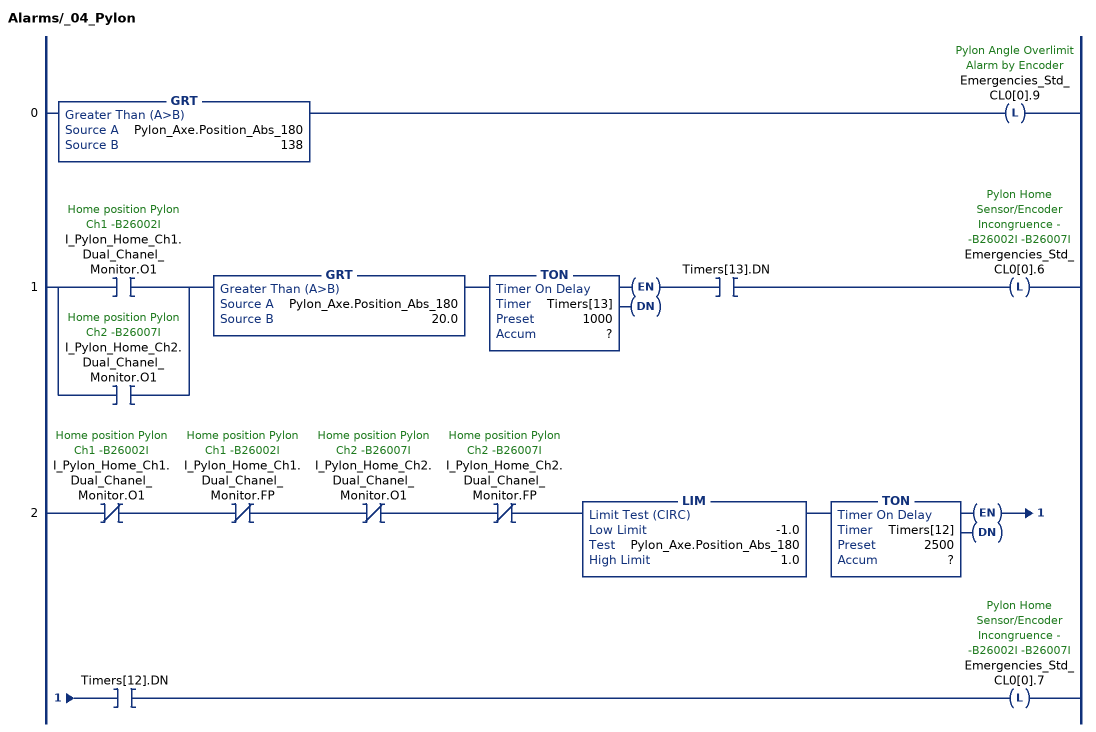
   0: GRT(Pylon_Axe.Position_Abs_180,138)OTL(Emergencies_Std_CL0[0].9);
   1: [XIC(I_Pylon_Home_Ch1.Dual_Chanel_Monitor.O1) ,XIC(I_Pylon_Home_Ch2.Dual_Chanel_Monitor.O1) ]GRT(Pylon_Axe.Position_Abs_180,20.0)TON(Timers[13],?,?)XIC(Timers[13].DN)OTL(Emergencies_Std_CL0[0].6);
   2: XIO(I_Pylon_Home_Ch1.Dual_Chanel_Monitor.O1)XIO(I_Pylon_Home_Ch1.Dual_Chanel_Monitor.FP)XIO(I_Pylon_Home_Ch2.Dual_Chanel_Monitor.O1)XIO(I_Pylon_Home_Ch2.Dual_Chanel_Monitor.FP)LIM(-1.0,Pylon_Axe.Position_Abs_180,1.0)TON(Timers[12],?,?)XIC(Timers[12].DN)OTL(Emergencies_Std_CL0[0].7);
END_ROUTINE

ROUTINE Main   (* ladder *)
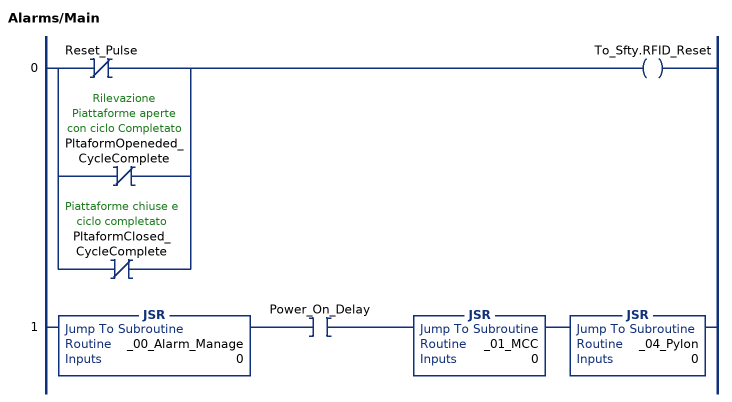
   0: [XIO(Reset_Pulse) ,XIO(PltaformOpeneded_CycleComplete) ,XIO(PltaformClosed_CycleComplete) ]OTE(To_Sfty.RFID_Reset);
   1: JSR(_00_Alarm_Manage,0)XIC(Power_On_Delay)JSR(_01_MCC,0)JSR(_04_Pylon,0);
END_ROUTINE
END_PROGRAM

PROGRAM General   (* main routine Main *)
VAR
   Avg_TimeInStation_CurrentHour : DINT := 303;
   Avg_TimeInStation_Daily : DINT := 207;
   Closing_CyclePlatTimes : DINT[20] := ([1] := 60000, [2] := 679, [3] := 679, [4] := 17399, [5] := 19639, [6] := 19639, [9] := 16239, [10] := 3400);
        [14]   // daily avg overall
        [13]   // daily total overall
        [11]   // daily total time waiting
        [10]   // Time Waiting on Lever,etc
        [9]   // Time Platform Move In Close
        [12]   // daily avg time waiting
   Cycle_Before_Timer : TIMER := (PRE := 60000);
   CyclePlatClose_Count_Daily : COUNTER := (PRE := 500);
   CyclePlatOpen_Count_Daily : COUNTER := (PRE := 500);
   DAY : DINT := 1;   // Day
   HMI_LapBars_Status : DINT := 1;   // 0 = Closed 1 = Opened 2 = Closing 3 = Opening
   HMI_Platform_Status : DINT := 1;   // 0 = Stopped 1 = Closing 2 = Closed 3 = Opening 4 = Opened
   HMI_reset_Partial_Life_Cycle : BOOL;
   HMI_reset_Partial_Life_RunHH : BOOL;
   HOUR : DINT := 19;   // Hour
   JM_Statistics_Hist : Run_Count_Hist_JM[100] := ([0].date[0] := 25, [0].date[1] := 11, [0].date[2] := 29, [0].runs[0] := 11, [0].runs[7] := 1, [0].runs[8] := 2, [0].runs[9] := 2, [0].runs[13] := 4, [0].runs[15] := 1, [0].runs[19] := 3, [0].time_avg[0] := 207, [0].time_avg[4] := 19639, [0].time_avg[5] := 22361, [0].time_avg[8] := 48, [0].time_avg[9] := 48, [0].time_avg[13] := 196, [0].time_avg[19] := 303, [1].date[0] := 25, [1].date[1] := 11, [1].date[2] := 28, [1].runs[0] := 65, [1].runs[8] := 2, [1].runs[9] := 1, [1].runs[15] := 3, [1].runs[16] := 7, [1].runs[17] := 8, [1].runs[18] := 8, [1].runs[19] := 8, [1].runs[20] := 8, [1].runs[21] := 7, [1].runs[22] := 8, [1].runs[23] := 5, [1].time_avg[0] := 204, [1].time_avg[2] := 3400, [1].time_avg[4] := 19639, [1].time_avg[5] := 22361, [1].time_avg[8] := 50, [1].time_avg[15] := 203, [1].time_avg[16] := 254, [1].time_avg[17] := 210, [1].time_avg[18] := 202, [1].time_avg[19] := 195, [1].time_avg[20] := 206, [1].time_avg[21] := 190, [1].time_avg[22] := 211, [1].time_avg[23] := 177, [2].date[0] := 25, [2].date[1] := 11, [2].date[2] := 27, [2].runs[0] := 63, [2].runs[14] := 6, [2].runs[15] := 4, [2].runs[16] := 7, [2].runs[17] := 7, [2].runs[18] := 8, [2].runs[19] := 8, [2].runs[20] := 7, [2].runs[21] := 5, [2].runs[22] := 8, [2].runs[23] := 3,
        [2].time_avg[0] := 234, [2].time_avg[4] := 21760, [2].time_avg[5] := 22361, [2].time_avg[14] := 167, [2].time_avg[15] := 316, [2].time_avg[16] := 272, [2].time_avg[17] := 206, [2].time_avg[18] := 208, [2].time_avg[19] := 242, [2].time_avg[20] := 266, [2].time_avg[21] := 233, [2].time_avg[22] := 223, [2].time_avg[23] := 245, [3].date[0] := 25, [3].date[1] := 11, [3].date[2] := 26, [3].runs[0] := 57, [3].runs[12] := 4, [3].runs[13] := 1, [3].runs[15] := 2, [3].runs[16] := 6, [3].runs[17] := 7, [3].runs[18] := 7, [3].runs[19] := 7, [3].runs[20] := 7, [3].runs[21] := 7, [3].runs[22] := 6, [3].runs[23] := 3, [3].time_avg[0] := 274, [3].time_avg[2] := 6041, [3].time_avg[4] := 21760, [3].time_avg[5] := 22361, [3].time_avg[12] := 396, [3].time_avg[13] := 320, [3].time_avg[15] := 271, [3].time_avg[16] := 271, [3].time_avg[17] := 292, [3].time_avg[18] := 243, [3].time_avg[19] := 255, [3].time_avg[20] := 243, [3].time_avg[21] := 289, [3].time_avg[22] := 278, [3].time_avg[23] := 283, [4].date[0] := 25, [4].date[1] := 11, [4].date[2] := 25, [4].runs[0] := 53, [4].runs[7] := 1, [4].runs[15] := 1, [4].runs[16] := 5, [4].runs[17] := 8, [4].runs[18] := 6, [4].runs[19] := 8, [4].runs[20] := 7, [4].runs[21] := 7, [4].runs[22] := 7, [4].runs[23] := 3, [4].time_avg[0] := 260, [4].time_avg[4] := 53080, [4].time_avg[5] := 22361,
        [4].time_avg[16] := 223, [4].time_avg[17] := 286, [4].time_avg[18] := 280, [4].time_avg[19] := 258, [4].time_avg[20] := 261, [4].time_avg[21] := 234, [4].time_avg[22] := 267, [4].time_avg[23] := 254, [5].date[0] := 25, [5].date[1] := 11, [5].date[2] := 24, [5].runs[0] := 67, [5].runs[7] := 4, [5].runs[8] := 3, [5].runs[10] := 2, [5].runs[11] := 4, [5].runs[13] := 1, [5].runs[14] := 1, [5].runs[15] := 4, [5].runs[16] := 7, [5].runs[17] := 7, [5].runs[18] := 7, [5].runs[19] := 7, [5].runs[20] := 4, [5].runs[21] := 7, [5].runs[22] := 6, [5].runs[23] := 3, [5].time_avg[0] := 254, [5].time_avg[2] := 76642, [5].time_avg[4] := 53080, [5].time_avg[5] := 22361, [5].time_avg[7] := 75, [5].time_avg[8] := 246, [5].time_avg[11] := 171, [5].time_avg[14] := 83, [5].time_avg[15] := 147, [5].time_avg[16] := 272, [5].time_avg[17] := 276, [5].time_avg[18] := 244, [5].time_avg[19] := 256, [5].time_avg[20] := 266, [5].time_avg[21] := 291, [5].time_avg[22] := 291, [5].time_avg[23] := 290, [6].date[0] := 25, [6].date[1] := 11, [6].date[2] := 23, [6].runs[0] := 54, [6].runs[10] := 2, [6].runs[11] := 4, [6].runs[15] := 1, [6].runs[16] := 8, [6].runs[17] := 7, [6].runs[18] := 6, [6].runs[19] := 5, [6].runs[20] := 8, [6].runs[21] := 6, [6].runs[22] := 5, [6].runs[23] := 2, [6].time_avg[0] := 268,
        [6].time_avg[4] := 23760, [6].time_avg[5] := 22361, [6].time_avg[11] := 332, [6].time_avg[16] := 211, [6].time_avg[17] := 253, [6].time_avg[18] := 262, [6].time_avg[19] := 274, [6].time_avg[20] := 241, [6].time_avg[21] := 295, [6].time_avg[22] := 310, [6].time_avg[23] := 371, [7].date[0] := 25, [7].date[1] := 11, [7].date[2] := 22, [7].runs[0] := 49, [7].runs[12] := 7, [7].runs[14] := 1, [7].runs[15] := 4, [7].runs[16] := 7, [7].runs[17] := 7, [7].runs[18] := 7, [7].runs[19] := 1, [7].runs[20] := 6, [7].runs[21] := 2, [7].runs[22] := 6, [7].runs[23] := 1, [7].time_avg[0] := 278, [7].time_avg[4] := 23760, [7].time_avg[5] := 22361, [7].time_avg[12] := 180, [7].time_avg[15] := 308, [7].time_avg[16] := 282, [7].time_avg[17] := 261, [7].time_avg[18] := 280, [7].time_avg[19] := 295, [7].time_avg[20] := 361, [7].time_avg[22] := 287, [8].date[0] := 25, [8].date[1] := 11, [8].date[2] := 20, [8].runs[0] := 58, [8].runs[10] := 2, [8].runs[11] := 3, [8].runs[13] := 5, [8].runs[14] := 4, [8].runs[15] := 3, [8].runs[16] := 5, [8].runs[17] := 4, [8].runs[18] := 3, [8].runs[19] := 6, [8].runs[20] := 5, [8].runs[21] := 7, [8].runs[22] := 7, [8].runs[23] := 4, [8].time_avg[0] := 205, [8].time_avg[2] := 15381, [8].time_avg[4] := 23760, [8].time_avg[5] := 22361, [8].time_avg[10] := 76, [8].time_avg[11] := 152,
        [8].time_avg[13] := 198, [8].time_avg[14] := 60, [8].time_avg[15] := 73, [8].time_avg[16] := 76, [8].time_avg[17] := 183, [8].time_avg[18] := 376, [8].time_avg[19] := 286, [8].time_avg[20] := 250, [8].time_avg[21] := 218, [8].time_avg[22] := 239, [8].time_avg[23] := 211, [9].date[0] := 25, [9].date[1] := 11, [9].date[2] := 19, [9].runs[0] := 7, [9].runs[12] := 2, [9].runs[13] := 4, [9].runs[17] := 1, [9].runs[18] := 1, [9].time_avg[0] := 217, [9].time_avg[2] := 78801, [9].time_avg[4] := 48480, [9].time_avg[5] := 22361, [9].time_avg[13] := 217, [10].date[0] := 25, [10].date[1] := 11, [10].date[2] := 16, [10].runs[0] := 7, [10].runs[10] := 2, [10].runs[13] := 7, [10].time_avg[0] := 93, [10].time_avg[4] := 27759, [10].time_avg[5] := 22361, [10].time_avg[13] := 93, [11].date[0] := 25, [11].date[1] := 11, [11].date[2] := 14, [11].runs[0] := 2, [11].runs[15] := 1, [11].runs[16] := 1, [11].time_avg[2] := 32760, [11].time_avg[4] := 27759, [11].time_avg[5] := 22361, [12].date[0] := 25, [12].date[1] := 11, [12].date[2] := 13, [12].runs[0] := 14, [12].runs[10] := 2, [12].runs[11] := 1, [12].runs[12] := 1, [12].runs[14] := 2, [12].runs[15] := 5, [12].runs[16] := 4, [12].runs[17] := 5, [12].time_avg[0] := 141, [12].time_avg[4] := 36240, [12].time_avg[5] := 22361, [12].time_avg[10] := 210, [12].time_avg[14] := 205, [12].time_avg[15] := 160,
        [12].time_avg[16] := 100, [12].time_avg[17] := 100, [13].date[0] := 25, [13].date[1] := 11, [13].date[2] := 11, [13].runs[0] := 2, [13].runs[18] := 2, [13].time_avg[0] := 88, [13].time_avg[4] := 36240, [13].time_avg[5] := 22361, [13].time_avg[18] := 88, [14].date[0] := 25, [14].date[1] := 11, [14].date[2] := 7, [14].runs[0] := 5, [14].runs[15] := 3, [14].runs[16] := 2, [14].time_avg[0] := 229, [14].time_avg[4] := 36240, [14].time_avg[5] := 22361, [14].time_avg[15] := 300, [14].time_avg[16] := 87, [15].date[0] := 25, [15].date[1] := 11, [15].date[2] := 6, [15].runs[0] := 13, [15].runs[15] := 1, [15].runs[16] := 3, [15].runs[17] := 8, [15].runs[18] := 1, [15].runs[19] := 4, [15].time_avg[0] := 54, [15].time_avg[4] := 36240, [15].time_avg[5] := 22361, [15].time_avg[17] := 46, [15].time_avg[19] := 66, [16].date[0] := 25, [16].date[1] := 10, [16].date[2] := 27, [16].runs[0] := 13, [16].runs[12] := 1, [16].runs[13] := 4, [16].runs[14] := 1, [16].time_avg[0] := 126, [16].time_avg[4] := 36240, [16].time_avg[5] := 22361, [16].time_avg[13] := 65, [17].date[0] := 25, [17].date[1] := 10, [17].date[2] := 26, [17].runs[0] := 58, [17].runs[10] := 1, [17].runs[11] := 2, [17].runs[12] := 3, [17].runs[13] := 8, [17].runs[14] := 8, [17].runs[15] := 6, [17].runs[16] := 7, [17].runs[17] := 7, [17].runs[18] := 6,
        [17].runs[19] := 7, [17].runs[20] := 3, [17].time_avg[0] := 252, [17].time_avg[2] := 40720, [17].time_avg[4] := 36240, [17].time_avg[5] := 22361, [17].time_avg[11] := 476, [17].time_avg[12] := 190, [17].time_avg[13] := 206, [17].time_avg[14] := 216, [17].time_avg[15] := 310, [17].time_avg[16] := 261, [17].time_avg[17] := 248, [17].time_avg[18] := 232, [17].time_avg[19] := 304, [17].time_avg[20] := 214, [18].date[0] := 25, [18].date[1] := 10, [18].date[2] := 25, [18].runs[0] := 47, [18].runs[12] := 5, [18].runs[13] := 9, [18].runs[14] := 5, [18].runs[16] := 2, [18].runs[17] := 8, [18].runs[18] := 7, [18].runs[19] := 7, [18].runs[20] := 4, [18].time_avg[0] := 227, [18].time_avg[4] := 26040, [18].time_avg[5] := 22361, [18].time_avg[12] := 203, [18].time_avg[13] := 166, [18].time_avg[14] := 231, [18].time_avg[16] := 370, [18].time_avg[17] := 239, [18].time_avg[18] := 252, [18].time_avg[19] := 244, [18].time_avg[20] := 235, [19].date[0] := 25, [19].date[1] := 10, [19].date[2] := 23, [19].runs[0] := 48, [19].runs[9] := 2, [19].runs[10] := 3, [19].runs[12] := 3, [19].runs[13] := 7, [19].runs[14] := 7, [19].runs[15] := 5, [19].runs[16] := 8, [19].runs[17] := 5, [19].runs[19] := 5, [19].runs[20] := 3, [19].time_avg[0] := 257, [19].time_avg[2] := 18201, [19].time_avg[4] := 26040, [19].time_avg[5] := 22361, [19].time_avg[9] := 102, [19].time_avg[10] := 259, [19].time_avg[12] := 493,
        [19].time_avg[13] := 241, [19].time_avg[14] := 231, [19].time_avg[15] := 264, [19].time_avg[16] := 252, [19].time_avg[17] := 280, [19].time_avg[19] := 300, [19].time_avg[20] := 235, [20].date[0] := 25, [20].date[1] := 10, [20].date[2] := 22, [20].runs[0] := 62, [20].runs[10] := 4, [20].runs[12] := 2, [20].runs[13] := 9, [20].runs[14] := 7, [20].runs[15] := 7, [20].runs[16] := 7, [20].runs[17] := 7, [20].runs[18] := 8, [20].runs[19] := 8, [20].runs[20] := 3, [20].time_avg[0] := 226, [20].time_avg[4] := 26079, [20].time_avg[5] := 22361, [20].time_avg[10] := 123, [20].time_avg[13] := 199, [20].time_avg[14] := 230, [20].time_avg[15] := 230, [20].time_avg[16] := 312, [20].time_avg[17] := 253, [20].time_avg[18] := 219, [20].time_avg[19] := 200, [20].time_avg[20] := 206, [21].date[0] := 25, [21].date[1] := 10, [21].date[2] := 21, [21].runs[0] := 58, [21].runs[11] := 3, [21].runs[12] := 1, [21].runs[13] := 8, [21].runs[14] := 7, [21].runs[15] := 4, [21].runs[16] := 8, [21].runs[17] := 8, [21].runs[18] := 7, [21].runs[19] := 8, [21].runs[20] := 4, [21].time_avg[0] := 233, [21].time_avg[2] := 42160, [21].time_avg[4] := 26079, [21].time_avg[5] := 22361, [21].time_avg[11] := 186, [21].time_avg[13] := 222, [21].time_avg[14] := 240, [21].time_avg[15] := 294, [21].time_avg[16] := 256, [21].time_avg[17] := 202, [21].time_avg[18] := 246, [21].time_avg[19] := 216, [21].time_avg[20] := 208,
        [22].date[0] := 25, [22].date[1] := 10, [22].date[2] := 20, [22].runs[0] := 47, [22].runs[10] := 2, [22].runs[11] := 6, [22].runs[12] := 1, [22].runs[13] := 7, [22].runs[14] := 7, [22].runs[15] := 7, [22].runs[16] := 4, [22].runs[17] := 1, [22].runs[18] := 2, [22].runs[19] := 7, [22].runs[20] := 3, [22].time_avg[0] := 249, [22].time_avg[2] := 52640, [22].time_avg[4] := 40960, [22].time_avg[5] := 22361, [22].time_avg[11] := 232, [22].time_avg[13] := 215, [22].time_avg[14] := 258, [22].time_avg[15] := 237, [22].time_avg[16] := 210, [22].time_avg[18] := 331, [22].time_avg[19] := 294, [22].time_avg[20] := 241, [23].date[0] := 25, [23].date[1] := 10, [23].date[2] := 19, [23].runs[0] := 61, [23].runs[9] := 2, [23].runs[10] := 2, [23].runs[11] := 8, [23].runs[12] := 4, [23].runs[13] := 6, [23].runs[14] := 1, [23].runs[15] := 8, [23].runs[16] := 7, [23].runs[17] := 7, [23].runs[18] := 7, [23].runs[19] := 7, [23].runs[20] := 2, [23].time_avg[0] := 237, [23].time_avg[2] := 59762, [23].time_avg[4] := 52320, [23].time_avg[5] := 22361, [23].time_avg[9] := 89, [23].time_avg[11] := 203, [23].time_avg[12] := 193, [23].time_avg[13] := 194, [23].time_avg[15] := 243, [23].time_avg[16] := 238, [23].time_avg[17] := 251, [23].time_avg[18] := 268, [23].time_avg[19] := 280, [23].time_avg[20] := 287, [24].date[0] := 25, [24].date[1] := 10, [24].date[2] := 18,
        [24].runs[0] := 51, [24].runs[9] := 2, [24].runs[10] := 5, [24].runs[11] := 8, [24].runs[12] := 2, [24].runs[13] := 5, [24].runs[14] := 6, [24].runs[15] := 7, [24].runs[16] := 5, [24].runs[17] := 7, [24].runs[18] := 4, [24].time_avg[0] := 246, [24].time_avg[4] := 52360, [24].time_avg[5] := 22361, [24].time_avg[10] := 182, [24].time_avg[11] := 228, [24].time_avg[12] := 212, [24].time_avg[13] := 231, [24].time_avg[14] := 324, [24].time_avg[15] := 255, [24].time_avg[16] := 238, [24].time_avg[17] := 263, [24].time_avg[18] := 255, [25].date[0] := 25, [25].date[1] := 10, [25].date[2] := 15, [25].runs[0] := 89, [25].runs[10] := 4, [25].runs[11] := 4, [25].runs[12] := 7, [25].runs[13] := 6, [25].runs[14] := 8, [25].runs[15] := 6, [25].runs[16] := 7, [25].runs[17] := 6, [25].time_avg[0] := 251, [25].time_avg[2] := 50482, [25].time_avg[4] := 52360, [25].time_avg[5] := 22361, [25].time_avg[10] := 61, [25].time_avg[11] := 214, [25].time_avg[12] := 261, [25].time_avg[13] := 348, [25].time_avg[14] := 197, [25].time_avg[15] := 264, [25].time_avg[16] := 241, [25].time_avg[17] := 309, [26].date[0] := 25, [26].date[1] := 10, [26].date[2] := 14, [26].runs[0] := 14, [26].runs[10] := 5, [26].runs[11] := 1, [26].runs[12] := 8, [26].time_avg[0] := 175, [26].time_avg[4] := 34119, [26].time_avg[5] := 22361, [26].time_avg[10] := 270, [26].time_avg[12] := 121, [27].date[0] := 25,
        [27].date[1] := 10, [27].date[2] := 13, [27].runs[0] := 29, [27].runs[12] := 3, [27].runs[13] := 5, [27].runs[14] := 6, [27].runs[15] := 4, [27].runs[16] := 7, [27].runs[17] := 4, [27].time_avg[0] := 256, [27].time_avg[2] := 63880, [27].time_avg[4] := 34119, [27].time_avg[5] := 22361, [27].time_avg[12] := 68, [27].time_avg[13] := 218, [27].time_avg[14] := 246, [27].time_avg[15] := 367, [27].time_avg[16] := 315, [27].time_avg[17] := 255, [28].date[0] := 25, [28].date[1] := 10, [28].date[2] := 10, [28].runs[0] := 27, [28].runs[9] := 9, [28].runs[10] := 11, [28].runs[11] := 7, [28].time_avg[0] := 89, [28].time_avg[4] := 33481, [28].time_avg[5] := 22361, [28].time_avg[9] := 82, [28].time_avg[10] := 83, [28].time_avg[11] := 123, [29].date[0] := 25, [29].date[1] := 10, [29].date[2] := 8, [29].runs[0] := 76, [29].runs[9] := 9, [29].runs[10] := 11, [29].runs[11] := 8, [29].runs[12] := 10, [29].runs[13] := 11, [29].runs[14] := 7, [29].runs[15] := 7, [29].runs[16] := 3, [29].time_avg[0] := 100, [29].time_avg[4] := 33481, [29].time_avg[5] := 22361, [29].time_avg[9] := 47, [29].time_avg[10] := 77, [29].time_avg[11] := 96, [29].time_avg[12] := 96, [29].time_avg[13] := 82, [29].time_avg[14] := 70, [29].time_avg[15] := 221, [29].time_avg[16] := 56, [30].date[0] := 25, [30].date[1] := 10, [30].date[2] := 7, [30].runs[0] := 1, [30].runs[8] := 1,
        [30].time_avg[4] := 33481, [30].time_avg[5] := 22361, [31].date[0] := 25, [31].date[1] := 10, [31].date[2] := 6, [31].runs[0] := 3, [31].runs[12] := 3, [31].time_avg[0] := 51, [31].time_avg[4] := 33481, [31].time_avg[5] := 22361, [31].time_avg[12] := 51, [32].date[0] := 25, [32].date[1] := 10, [32].date[2] := 5, [32].runs[0] := 3, [32].runs[12] := 1, [32].runs[15] := 2, [32].time_avg[0] := 43, [32].time_avg[4] := 33481, [32].time_avg[5] := 22361, [32].time_avg[15] := 43, [33].date[0] := 25, [33].date[1] := 10, [33].date[2] := 4, [33].runs[0] := 15, [33].runs[10] := 4, [33].runs[11] := 3, [33].runs[12] := 3, [33].runs[15] := 4, [33].runs[16] := 1, [33].time_avg[0] := 228, [33].time_avg[2] := 47342, [33].time_avg[4] := 33481, [33].time_avg[5] := 22361, [33].time_avg[10] := 258, [33].time_avg[11] := 342, [33].time_avg[12] := 69, [33].time_avg[15] := 112, [34].date[0] := 25, [34].date[1] := 10, [34].date[2] := 1, [34].runs[0] := 64, [34].runs[9] := 1, [34].runs[10] := 7, [34].runs[11] := 8, [34].runs[12] := 9, [34].runs[13] := 6, [34].runs[14] := 8, [34].runs[15] := 9, [34].runs[16] := 8, [34].runs[17] := 8, [34].time_avg[0] := 168, [34].time_avg[4] := 53200, [34].time_avg[5] := 22361, [34].time_avg[10] := 151, [34].time_avg[11] := 172, [34].time_avg[12] := 168, [34].time_avg[13] := 171, [34].time_avg[14] := 150, [34].time_avg[15] := 177,
        [34].time_avg[16] := 175, [34].time_avg[17] := 175, [35].date[0] := 25, [35].date[1] := 9, [35].date[2] := 30, [35].runs[0] := 60, [35].runs[9] := 5, [35].runs[10] := 5, [35].runs[11] := 9, [35].runs[12] := 7, [35].runs[13] := 8, [35].runs[14] := 9, [35].runs[15] := 9, [35].runs[16] := 8, [35].time_avg[0] := 176, [35].time_avg[2] := 40561, [35].time_avg[4] := 53200, [35].time_avg[5] := 22361, [35].time_avg[9] := 120, [35].time_avg[10] := 150, [35].time_avg[11] := 176, [35].time_avg[12] := 186, [35].time_avg[13] := 219, [35].time_avg[14] := 153, [35].time_avg[15] := 180, [35].time_avg[16] := 165, [36].date[0] := 25, [36].date[1] := 9, [36].date[2] := 29, [36].runs[0] := 57, [36].runs[8] := 2, [36].runs[9] := 7, [36].runs[10] := 7, [36].runs[11] := 8, [36].runs[12] := 5, [36].runs[13] := 7, [36].runs[14] := 7, [36].runs[15] := 7, [36].runs[16] := 7, [36].time_avg[0] := 211, [36].time_avg[4] := 56839, [36].time_avg[5] := 22361, [36].time_avg[9] := 166, [36].time_avg[10] := 267, [36].time_avg[11] := 147, [36].time_avg[12] := 241, [36].time_avg[13] := 205, [36].time_avg[14] := 168, [36].time_avg[15] := 266, [36].time_avg[16] := 222, [37].date[0] := 25, [37].date[1] := 9, [37].date[2] := 28, [37].runs[0] := 58, [37].runs[9] := 3, [37].runs[10] := 9, [37].runs[11] := 7, [37].runs[12] := 8, [37].runs[13] := 8, [37].runs[14] := 8,
        [37].runs[15] := 7, [37].runs[16] := 8, [37].time_avg[0] := 184, [37].time_avg[4] := 56839, [37].time_avg[5] := 22361, [37].time_avg[9] := 167, [37].time_avg[10] := 193, [37].time_avg[11] := 208, [37].time_avg[12] := 169, [37].time_avg[13] := 199, [37].time_avg[14] := 199, [37].time_avg[15] := 173, [37].time_avg[16] := 151, [38].date[0] := 25, [38].date[1] := 9, [38].date[2] := 25, [38].runs[0] := 64, [38].runs[8] := 4, [38].runs[9] := 6, [38].runs[10] := 7, [38].runs[11] := 7, [38].runs[12] := 8, [38].runs[13] := 8, [38].runs[14] := 8, [38].runs[15] := 9, [38].runs[16] := 7, [38].time_avg[0] := 201, [38].time_avg[4] := 56839, [38].time_avg[5] := 22361, [38].time_avg[8] := 455, [38].time_avg[9] := 193, [38].time_avg[10] := 212, [38].time_avg[11] := 189, [38].time_avg[12] := 207, [38].time_avg[13] := 224, [38].time_avg[14] := 191, [38].time_avg[15] := 166, [38].time_avg[16] := 193, [39].date[0] := 25, [39].date[1] := 9, [39].date[2] := 24, [39].runs[0] := 50, [39].runs[9] := 4, [39].runs[10] := 6, [39].runs[11] := 5, [39].runs[12] := 6, [39].runs[13] := 5, [39].runs[14] := 8, [39].runs[15] := 8, [39].runs[16] := 8, [39].time_avg[0] := 195, [39].time_avg[4] := 56839, [39].time_avg[5] := 22361, [39].time_avg[9] := 83, [39].time_avg[10] := 198, [39].time_avg[11] := 260, [39].time_avg[12] := 133, [39].time_avg[13] := 207, [39].time_avg[14] := 244, [39].time_avg[15] := 215,
        [39].time_avg[16] := 169, [40].date[0] := 25, [40].date[1] := 9, [40].date[2] := 22, [40].runs[0] := 46, [40].runs[8] := 4, [40].runs[9] := 3, [40].runs[10] := 7, [40].runs[11] := 5, [40].runs[12] := 7, [40].runs[13] := 5, [40].runs[14] := 2, [40].runs[15] := 6, [40].runs[16] := 7, [40].time_avg[0] := 229, [40].time_avg[4] := 56839, [40].time_avg[5] := 22361, [40].time_avg[8] := 208, [40].time_avg[10] := 179, [40].time_avg[11] := 196, [40].time_avg[12] := 160, [40].time_avg[13] := 227, [40].time_avg[15] := 325, [40].time_avg[16] := 281, [41].date[0] := 25, [41].date[1] := 9, [41].date[2] := 21, [41].runs[0] := 9, [41].runs[8] := 1, [41].runs[9] := 6, [41].runs[14] := 2, [41].time_avg[0] := 233, [41].time_avg[2] := 43360, [41].time_avg[4] := 56839, [41].time_avg[5] := 22361, [41].time_avg[9] := 244, [41].time_avg[14] := 175, [42].date[0] := 25, [42].date[1] := 9, [42].date[2] := 18, [42].runs[0] := 6, [42].runs[11] := 5, [42].runs[12] := 1, [42].time_avg[0] := 226, [42].time_avg[4] := 37320, [42].time_avg[5] := 22361, [42].time_avg[11] := 226, [43].date[0] := 25, [43].date[1] := 9, [43].date[2] := 16, [43].runs[0] := 2, [43].runs[15] := 1, [43].runs[16] := 1, [43].time_avg[2] := 46801, [43].time_avg[4] := 37320, [43].time_avg[5] := 22361, [44].date[0] := 25, [44].date[1] := 8, [44].date[2] := 15, [44].runs[0] := 3,
        [44].runs[12] := 1, [44].runs[15] := 2, [44].time_avg[4] := 37641, [44].time_avg[5] := 22361, [45].date[0] := 25, [45].date[1] := 7, [45].date[2] := 13, [45].runs[0] := 107, [45].runs[9] := 2, [45].runs[14] := 2, [45].runs[16] := 8, [45].time_avg[0] := 162, [45].time_avg[2] := 22208, [45].time_avg[4] := 37641, [45].time_avg[5] := 22361, [45].time_avg[9] := 55, [45].time_avg[14] := 220, [45].time_avg[16] := 142, [46].date[0] := -2, [46].date[1] := 1, [46].date[2] := 15, [46].runs[0] := 1, [46].time_avg[4] := 45599, [46].time_avg[5] := 22361, [47].date[0] := -2, [47].date[1] := 1, [47].date[2] := 12, [47].runs[0] := 14, [47].runs[23] := 3, [47].time_avg[0] := 172, [47].time_avg[4] := 45599, [47].time_avg[5] := 22361, [47].time_avg[23] := 108, [48].date[0] := -2, [48].date[1] := 1, [48].date[2] := 11, [48].runs[0] := 14, [48].runs[21] := 1, [48].time_avg[0] := 145, [48].time_avg[4] := 45599, [48].time_avg[5] := 22361, [49].date[0] := -2, [49].date[1] := 1, [49].date[2] := 10, [49].runs[0] := 2, [49].runs[20] := 1, [49].runs[23] := 1, [49].time_avg[4] := 45599, [49].time_avg[5] := 22361, [50].date[0] := -2, [50].date[1] := 1, [50].date[2] := 8, [50].runs[0] := 1, [50].time_avg[4] := 45599, [50].time_avg[5] := 22361, [51].date[0] := -2, [51].date[1] := 1, [51].date[2] := 6, [51].runs[0] := 2, [51].runs[20] := 1,
        [51].time_avg[4] := 45599, [51].time_avg[5] := 22361, [52].date[0] := -2, [52].date[1] := 1, [52].date[2] := 5, [52].runs[0] := 10, [52].runs[20] := 2, [52].runs[23] := 3, [52].time_avg[0] := 139, [52].time_avg[4] := 45599, [52].time_avg[5] := 22361, [52].time_avg[23] := 139, [53].date[0] := -2, [53].date[1] := 1, [53].date[2] := 4, [53].runs[0] := 7, [53].runs[21] := 1, [53].runs[22] := 2, [53].time_avg[0] := 542, [53].time_avg[4] := 45599, [53].time_avg[5] := 22361, [53].time_avg[22] := 542, [54].date[0] := -2, [54].date[1] := 1, [54].date[2] := 2, [54].runs[0] := 4, [54].runs[23] := 4, [54].time_avg[4] := 45599, [54].time_avg[5] := 22361, [55].date[0] := -2, [55].date[1] := 1, [55].date[2] := 21, [55].runs[0] := 12, [55].runs[19] := 1, [55].runs[20] := 1, [55].runs[23] := 2, [55].time_avg[0] := 325, [55].time_avg[4] := 45599, [55].time_avg[5] := 22361, [56].date[0] := -2, [56].date[1] := 1, [56].date[2] := 20, [56].runs[0] := 15, [56].runs[17] := 4, [56].runs[18] := 1, [56].runs[23] := 1, [56].time_avg[0] := 214, [56].time_avg[2] := 35440, [56].time_avg[4] := 45599, [56].time_avg[5] := 22361, [56].time_avg[17] := 368, [57].date[0] := -2, [57].date[1] := 1, [57].date[2] := 19, [57].runs[0] := 6, [57].runs[17] := 1, [57].runs[18] := 2, [57].time_avg[0] := 112, [57].time_avg[2] := 41643, [57].time_avg[4] := 46281,
        [57].time_avg[5] := 22361, [57].time_avg[18] := 87, [58].date[0] := -2, [58].date[1] := 1, [58].date[2] := 15, [58].runs[0] := 7, [58].time_avg[0] := 126, [58].time_avg[4] := 37560, [58].time_avg[5] := 22361, [59].date[0] := -2, [59].date[1] := 1, [59].date[2] := 13, [59].runs[0] := 32, [59].runs[20] := 8, [59].runs[21] := 5, [59].runs[23] := 6, [59].time_avg[0] := 213, [59].time_avg[4] := 37560, [59].time_avg[5] := 22361, [59].time_avg[20] := 70, [59].time_avg[21] := 68, [59].time_avg[23] := 68, [60].date[0] := -2, [60].date[1] := 1, [60].date[2] := 12, [60].runs[0] := 17, [60].runs[20] := 5, [60].runs[21] := 5, [60].time_avg[0] := 121, [60].time_avg[4] := 37560, [60].time_avg[5] := 22361, [60].time_avg[20] := 167, [60].time_avg[21] := 64, [61].date[0] := -2, [61].date[1] := 1, [61].date[2] := 11, [61].runs[0] := 8, [61].runs[18] := 1, [61].runs[19] := 2, [61].runs[20] := 2, [61].runs[23] := 3, [61].time_avg[0] := 204, [61].time_avg[4] := 37560, [61].time_avg[5] := 22361, [61].time_avg[19] := 278, [61].time_avg[23] := 58, [62].date[0] := -2, [62].date[1] := 1, [62].date[2] := 10, [62].runs[0] := 4, [62].runs[18] := 1, [62].runs[20] := 2, [62].runs[23] := 1, [62].time_avg[0] := 4, [62].time_avg[2] := 30360, [62].time_avg[4] := 37560, [62].time_avg[5] := 22361, [62].time_avg[20] := 317, [63].date[0] := -2, [63].date[1] := 1,
        [63].date[2] := 8, [63].runs[0] := 28, [63].runs[17] := 1, [63].runs[18] := 1, [63].runs[20] := 4, [63].runs[21] := 2, [63].runs[23] := 3, [63].time_avg[0] := 184, [63].time_avg[2] := -4678, [63].time_avg[4] := 9800, [63].time_avg[5] := 22361, [63].time_avg[18] := 298, [63].time_avg[20] := 114, [63].time_avg[23] := 244, [64].date[0] := -2, [64].date[1] := 1, [64].date[2] := 7, [64].runs[0] := 9, [64].runs[17] := 1, [64].runs[19] := 1, [64].runs[20] := 3, [64].time_avg[0] := 370, [64].time_avg[5] := 22361, [64].time_avg[20] := 370, [65].date[0] := -2, [65].date[1] := 2, [65].date[2] := 10, [65].runs[0] := 14, [65].runs[19] := 9, [65].runs[20] := 5, [65].time_avg[5] := 22361, [66].date[0] := 20, [66].date[1] := 3, [66].date[2] := 5, [66].runs[0] := 11, [66].runs[8] := 1, [66].runs[9] := 1, [66].runs[10] := 1, [66].runs[14] := 3, [66].runs[15] := 1, [66].runs[16] := 2, [66].runs[17] := 2, [66].time_avg[0] := 250, [66].time_avg[5] := 22361, [66].time_avg[10] := 454, [66].time_avg[14] := 139, [66].time_avg[16] := 157, [67].date[0] := 20, [67].date[1] := 3, [67].date[2] := 4, [67].runs[0] := 20, [67].runs[11] := 4, [67].runs[12] := 6, [67].runs[18] := 8, [67].runs[19] := 2, [67].time_avg[0] := 36, [67].time_avg[2] := 31218, [67].time_avg[5] := 22361, [67].time_avg[12] := 36, [68].date[0] := 20,
        [68].date[1] := 3, [68].date[2] := 2, [68].runs[0] := 87, [68].runs[12] := 1, [68].runs[13] := 6, [68].runs[14] := 17, [68].runs[15] := 16, [68].runs[16] := 15, [68].runs[17] := 15, [68].runs[18] := 11, [68].runs[19] := 6, [68].time_avg[0] := 29, [68].time_avg[4] := 28480, [68].time_avg[5] := 22361, [68].time_avg[14] := 29, [68].time_avg[15] := 23, [68].time_avg[16] := 34, [68].time_avg[17] := 29, [68].time_avg[18] := 26, [69].date[0] := -2, [69].date[1] := 1, [69].date[2] := 11, [69].runs[0] := 114, [69].runs[7] := 7, [69].runs[9] := 2, [69].runs[10] := 8, [69].runs[11] := 3, [69].runs[13] := 6, [69].runs[14] := 11, [69].time_avg[0] := 84, [69].time_avg[2] := 22683, [69].time_avg[4] := 28480, [69].time_avg[5] := 22361, [69].time_avg[7] := 107, [69].time_avg[11] := 24, [69].time_avg[13] := 70, [69].time_avg[14] := 104, [70].date[0] := -2, [70].date[1] := 1, [70].date[2] := 8, [70].runs[0] := 19, [70].runs[23] := 3, [70].time_avg[0] := 35, [70].time_avg[4] := 23240, [70].time_avg[5] := 22361, [71].date[0] := -2, [71].date[1] := 1, [71].date[2] := 7, [71].runs[0] := 30, [71].runs[20] := 2, [71].runs[21] := 6, [71].runs[22] := 1, [71].time_avg[0] := 199, [71].time_avg[4] := 23240, [71].time_avg[5] := 22361, [71].time_avg[21] := 199, [72].date[0] := -2, [72].date[1] := 1, [72].date[2] := 6, [72].runs[0] := 30,
        [72].time_avg[4] := 23240, [72].time_avg[5] := 22361, [73].date[0] := -2, [73].date[1] := 1, [73].date[2] := 5, [73].runs[0] := 4, [73].runs[23] := 1, [73].time_avg[4] := 23240, [73].time_avg[5] := 22361, [74].date[0] := 19, [74].date[1] := 9, [74].date[2] := 3, [74].runs[0] := 62, [74].runs[7] := 1, [74].runs[9] := 3, [74].runs[10] := 4, [74].runs[11] := 7, [74].runs[12] := 7, [74].runs[13] := 9, [74].runs[14] := 7, [74].runs[15] := 8, [74].runs[16] := 7, [74].runs[17] := 8, [74].runs[18] := 1, [74].runs[21] := 1, [74].time_avg[0] := 211, [74].time_avg[2] := 5236, [74].time_avg[3] := 12461, [74].time_avg[4] := 23240, [74].time_avg[5] := 22361, [74].time_avg[12] := 175, [74].time_avg[13] := 206, [74].time_avg[17] := 252, [74].time_avg[18] := 206, [74].time_avg[21] := 206, [75].date[0] := 19, [75].date[1] := 9, [75].date[2] := 2, [75].runs[0] := 70, [75].runs[7] := 1, [75].runs[9] := 4, [75].runs[10] := 3, [75].runs[12] := 6, [75].runs[13] := 7, [75].runs[14] := 5, [75].runs[15] := 9, [75].runs[16] := 7, [75].runs[17] := 2, [75].runs[18] := 8, [75].runs[19] := 9, [75].runs[20] := 8, [75].runs[21] := 1, [75].time_avg[0] := 186, [75].time_avg[2] := 5622, [75].time_avg[3] := 14544, [75].time_avg[4] := 20279, [75].time_avg[5] := 21563, [75].time_avg[10] := 214, [75].time_avg[12] := 152, [75].time_avg[13] := 173,
        [75].time_avg[14] := 183, [75].time_avg[15] := 191, [75].time_avg[16] := 193, [75].time_avg[17] := 150, [75].time_avg[18] := 177, [75].time_avg[19] := 190, [75].time_avg[20] := 190, [75].time_avg[21] := 370, [76].date[0] := 19, [76].date[1] := 9, [76].date[2] := 1, [76].runs[0] := 118, [76].runs[7] := 1, [76].runs[8] := 4, [76].runs[9] := 9, [76].runs[10] := 8, [76].runs[11] := 8, [76].runs[12] := 7, [76].runs[13] := 5, [76].runs[14] := 8, [76].runs[15] := 8, [76].runs[16] := 9, [76].runs[17] := 8, [76].runs[18] := 8, [76].runs[19] := 8, [76].runs[20] := 11, [76].runs[21] := 9, [76].runs[22] := 7, [76].time_avg[0] := 197, [76].time_avg[2] := 7812, [76].time_avg[3] := 8907, [76].time_avg[4] := 17438, [76].time_avg[5] := 20839, [76].time_avg[11] := 228, [76].time_avg[12] := 233, [76].time_avg[15] := 183, [76].time_avg[16] := 195, [76].time_avg[17] := 218, [76].time_avg[18] := 219, [76].time_avg[19] := 279, [76].time_avg[20] := 132, [76].time_avg[21] := 181, [76].time_avg[22] := 154, [77].date[0] := 19, [77].date[1] := 8, [77].date[2] := 31, [77].runs[0] := 121, [77].runs[7] := 1, [77].runs[9] := 6, [77].runs[10] := 11, [77].runs[11] := 8, [77].runs[12] := 9, [77].runs[13] := 9, [77].runs[14] := 9, [77].runs[15] := 8, [77].runs[16] := 9, [77].runs[17] := 9, [77].runs[18] := 9, [77].runs[19] := 9, [77].runs[20] := 10,
        [77].runs[21] := 8, [77].runs[22] := 6, [77].time_avg[0] := 193, [77].time_avg[2] := 4893, [77].time_avg[3] := 10185, [77].time_avg[4] := 20961, [77].time_avg[5] := 18600, [77].time_avg[10] := 199, [77].time_avg[11] := 202, [77].time_avg[12] := 189, [77].time_avg[13] := 205, [77].time_avg[14] := 168, [77].time_avg[15] := 213, [77].time_avg[16] := 188, [77].time_avg[17] := 210, [77].time_avg[18] := 201, [77].time_avg[19] := 185, [77].time_avg[20] := 174, [77].time_avg[21] := 198, [77].time_avg[22] := 164, [78].date[0] := 19, [78].date[1] := 8, [78].date[2] := 30, [78].runs[0] := 102, [78].runs[7] := 1, [78].runs[9] := 4, [78].runs[10] := 4, [78].runs[11] := 8, [78].runs[12] := 9, [78].runs[13] := 8, [78].runs[14] := 8, [78].runs[15] := 9, [78].runs[16] := 8, [78].runs[17] := 7, [78].runs[18] := 6, [78].runs[19] := 9, [78].runs[20] := 9, [78].runs[21] := 8, [78].runs[22] := 4, [78].time_avg[0] := 212, [78].time_avg[2] := 6981, [78].time_avg[3] := 13438, [78].time_avg[4] := 22920, [78].time_avg[5] := 22402, [78].time_avg[11] := 206, [78].time_avg[12] := 233, [78].time_avg[13] := 225, [78].time_avg[14] := 202, [78].time_avg[15] := 222, [78].time_avg[16] := 214, [78].time_avg[17] := 168, [78].time_avg[18] := 226, [78].time_avg[19] := 184, [78].time_avg[20] := 240, [78].time_avg[21] := 205, [78].time_avg[22] := 200, [79].date[0] := 19, [79].date[1] := 8, [79].date[2] := 29, [79].runs[0] := 108,
        [79].runs[9] := 4, [79].runs[10] := 5, [79].runs[11] := 9, [79].runs[12] := 10, [79].runs[13] := 10, [79].runs[14] := 10, [79].runs[15] := 8, [79].runs[16] := 9, [79].runs[17] := 10, [79].runs[18] := 9, [79].runs[19] := 9, [79].runs[20] := 9, [79].runs[21] := 5, [79].time_avg[0] := 182, [79].time_avg[2] := 4017, [79].time_avg[3] := 9797, [79].time_avg[4] := 23082, [79].time_avg[5] := 18998, [79].time_avg[10] := 174, [79].time_avg[11] := 200, [79].time_avg[12] := 157, [79].time_avg[13] := 156, [79].time_avg[14] := 151, [79].time_avg[15] := 216, [79].time_avg[16] := 184, [79].time_avg[17] := 179, [79].time_avg[18] := 206, [79].time_avg[19] := 187, [79].time_avg[20] := 186, [79].time_avg[21] := 214, [80].date[0] := 19, [80].date[1] := 8, [80].date[2] := 28, [80].runs[0] := 107, [80].runs[7] := 2, [80].runs[8] := 5, [80].runs[9] := 11, [80].runs[10] := 6, [80].runs[11] := 9, [80].runs[12] := 9, [80].runs[13] := 10, [80].runs[14] := 9, [80].runs[15] := 7, [80].runs[16] := 9, [80].runs[17] := 9, [80].runs[18] := 8, [80].runs[19] := 9, [80].runs[20] := 8, [80].runs[21] := 1, [80].time_avg[0] := 204, [80].time_avg[2] := 4432, [80].time_avg[3] := 11019, [80].time_avg[4] := 18000, [80].time_avg[5] := 22000, [80].time_avg[10] := 191, [80].time_avg[11] := 184, [80].time_avg[12] := 190, [80].time_avg[13] := 174, [80].time_avg[14] := 198, [80].time_avg[15] := 270,
        [80].time_avg[16] := 203, [80].time_avg[17] := 194, [80].time_avg[18] := 256, [80].time_avg[19] := 195, [80].time_avg[20] := 206, [80].time_avg[21] := 186, [81].date[0] := 19, [81].date[1] := 8, [81].date[2] := 27, [81].runs[0] := 114, [81].runs[7] := 1, [81].runs[9] := 4, [81].runs[10] := 5, [81].runs[11] := 9, [81].runs[12] := 8, [81].runs[13] := 8, [81].runs[14] := 9, [81].runs[15] := 11, [81].runs[16] := 10, [81].runs[17] := 11, [81].runs[18] := 11, [81].runs[19] := 12, [81].runs[20] := 9, [81].runs[21] := 6, [81].time_avg[0] := 146, [81].time_avg[2] := 5205, [81].time_avg[3] := 8324, [81].time_avg[4] := 51040, [81].time_avg[5] := 27563, [81].time_avg[10] := 152, [81].time_avg[11] := 179, [81].time_avg[12] := 150, [81].time_avg[13] := 187, [81].time_avg[14] := 179, [81].time_avg[15] := 142, [81].time_avg[16] := 146, [81].time_avg[17] := 112, [81].time_avg[18] := 141, [81].time_avg[19] := 93, [81].time_avg[20] := 163, [81].time_avg[21] := 149, [82].date[0] := 19, [82].date[1] := 8, [82].date[2] := 26, [82].runs[0] := 110, [82].runs[7] := 1, [82].runs[9] := 4, [82].runs[10] := 5, [82].runs[11] := 8, [82].runs[12] := 9, [82].runs[13] := 10, [82].runs[14] := 10, [82].runs[15] := 9, [82].runs[16] := 10, [82].runs[17] := 10, [82].runs[18] := 9, [82].runs[19] := 10, [82].runs[20] := 10, [82].runs[21] := 5, [82].time_avg[0] := 168,
        [82].time_avg[2] := 4284, [82].time_avg[3] := 14914, [82].time_avg[4] := 18760, [82].time_avg[5] := 19159, [82].time_avg[10] := 159, [82].time_avg[11] := 212, [82].time_avg[12] := 159, [82].time_avg[13] := 168, [82].time_avg[14] := 162, [82].time_avg[15] := 181, [82].time_avg[16] := 170, [82].time_avg[17] := 150, [82].time_avg[18] := 164, [82].time_avg[19] := 159, [82].time_avg[20] := 161, [82].time_avg[21] := 183, [83].date[0] := 19, [83].date[1] := 8, [83].date[2] := 25, [83].runs[0] := 116, [83].runs[7] := 1, [83].runs[9] := 4, [83].runs[10] := 4, [83].runs[11] := 9, [83].runs[12] := 9, [83].runs[13] := 9, [83].runs[14] := 11, [83].runs[15] := 10, [83].runs[16] := 9, [83].runs[17] := 9, [83].runs[18] := 7, [83].runs[19] := 11, [83].runs[20] := 9, [83].runs[21] := 10, [83].runs[22] := 4, [83].time_avg[0] := 171, [83].time_avg[2] := 3326, [83].time_avg[3] := 10694, [83].time_avg[4] := 30960, [83].time_avg[5] := 24322, [83].time_avg[10] := 258, [83].time_avg[11] := 206, [83].time_avg[12] := 166, [83].time_avg[13] := 166, [83].time_avg[14] := 133, [83].time_avg[15] := 149, [83].time_avg[16] := 187, [83].time_avg[17] := 204, [83].time_avg[18] := 204, [83].time_avg[19] := 143, [83].time_avg[20] := 164, [83].time_avg[21] := 145, [83].time_avg[22] := 212, [84].date[0] := 19, [84].date[1] := 8, [84].date[2] := 24, [84].runs[0] := 116, [84].runs[7] := 1, [84].runs[9] := 4, [84].runs[10] := 5,